   // stn[29].wipBtn[35,0] := 1000;
   // stn[29].wipBtn[35,1] := 1000;
   // stn[29].wipBtn[35,2] := 1000;
   // stn[29].wipBtn[35,3] := 1000;
   // stn[29].wipBtn[35,4] := 1000;
   // stn[29].wipBtn[35,5] := 1000;
   // stn[29].wipBtn[35,6] := 1000;
   // stn[29].wipBtn[35,7] := 1000;
   // stn[29].wipBtn[36,0] := 1000;
   // stn[29].wipBtn[36,1] := 1000;
   // stn[29].wipBtn[36,2] := 1000;
   // stn[29].wipBtn[36,3] := 1000;
   // stn[29].wipBtn[36,4] := 1000;
   // stn[29].wipBtn[36,5] := 1000;
   // stn[29].wipBtn[36,6] := 1000;
   // stn[29].wipBtn[36,7] := 1000;
   // stn[29].wipBtn[37,0] := 1000;
   // stn[29].wipBtn[37,1] := 1000;
   // stn[29].wipBtn[37,2] := 1000;
   // stn[29].wipBtn[37,3] := 1000;
   // stn[29].wipBtn[37,4] := 1000;
   // stn[29].wipBtn[37,5] := 1000;
   // stn[29].wipBtn[37,6] := 1000;
   // stn[29].wipBtn[37,7] := 1000;
   // stn[29].wipBtn[38,0] := 1000;
   // stn[29].wipBtn[38,1] := 1000;
   // stn[29].wipBtn[38,2] := 1000;
   // stn[29].wipBtn[38,3] := 1000;
   // stn[29].wipBtn[38,4] := 1000;
   // stn[29].wipBtn[38,5] := 1000;
   // stn[29].wipBtn[38,6] := 1000;
   // stn[29].wipBtn[38,7] := 1000;
   // stn[29].wipBtn[39,0] := 1000;
   // stn[29].wipBtn[39,1] := 1000;
   // stn[29].wipBtn[39,2] := 1000;
   // stn[29].wipBtn[39,3] := 1000;
   // stn[29].wipBtn[39,4] := 1000;
   // stn[29].wipBtn[39,5] := 1000;
   // stn[29].wipBtn[39,6] := 1000;
   // stn[29].wipBtn[39,7] := 1000;
   // stn[29].wipBtn[40,0] := 1000;
   // stn[29].wipBtn[40,1] := 1000;
   // stn[29].wipBtn[40,2] := 1000;
   // stn[29].wipBtn[40,3] := 1000;
   // stn[29].wipBtn[40,4] := 1000;
   // stn[29].wipBtn[40,5] := 1000;
   // stn[29].wipBtn[40,6] := 1000;
   // stn[29].wipBtn[40,7] := 1000;
   // stn[29].wipBtn[41,0] := 1000;
   // stn[29].wipBtn[41,1] := 1000;
   // stn[29].wipBtn[41,2] := 1000;
   // stn[29].wipBtn[41,3] := 1000;
   // stn[29].wipBtn[41,4] := 1000;
   // stn[29].wipBtn[41,5] := 1000;
   // stn[29].wipBtn[41,6] := 1000;
   // stn[29].wipBtn[41,7] := 1000;
   // stn[29].wipBtn[42,0] := 1000;
   // stn[29].wipBtn[42,1] := 1000;
   // stn[29].wipBtn[42,2] := 1000;
   // stn[29].wipBtn[42,3] := 1000;
   // stn[29].wipBtn[42,4] := 1000;
   // stn[29].wipBtn[42,5] := 1000;
   // stn[29].wipBtn[42,6] := 1000;
   // stn[29].wipBtn[42,7] := 1000;
   // stn[29].wipBtn[43,0] := 1000;
   // stn[29].wipBtn[43,1] := 1000;
   // stn[29].wipBtn[43,2] := 1000;
   // stn[29].wipBtn[43,3] := 1000;
   // stn[29].wipBtn[43,4] := 1000;
   // stn[29].wipBtn[43,5] := 1000;
   // stn[29].wipBtn[43,6] := 1000;
   // stn[29].wipBtn[43,7] := 1000;
   // stn[29].wipBtn[44,0] := 1000;
   // stn[29].wipBtn[44,1] := 1000;
   // stn[29].wipBtn[44,2] := 1000;
   // stn[29].wipBtn[44,3] := 1000;
   // stn[29].wipBtn[44,4] := 1000;
   // stn[29].wipBtn[44,5] := 1000;
   // stn[29].wipBtn[44,6] := 1000;
   // stn[29].wipBtn[44,7] := 1000;
   // stn[29].wipBtn[45,0] := 1000;
   // stn[29].wipBtn[45,1] := 1000;
   // stn[29].wipBtn[45,2] := 1000;
   // stn[29].wipBtn[45,3] := 1000;
   // stn[29].wipBtn[45,4] := 1000;
   // stn[29].wipBtn[45,5] := 1000;
   // stn[29].wipBtn[45,6] := 1000;
   // stn[29].wipBtn[45,7] := 1000;
   // stn[29].wipBtn[46,0] := 1000;
   // stn[29].wipBtn[46,1] := 1000;
   // stn[29].wipBtn[46,2] := 1000;
   // stn[29].wipBtn[46,3] := 1000;
   // stn[29].wipBtn[46,4] := 1000;
   // stn[29].wipBtn[46,5] := 1000;
   // stn[29].wipBtn[46,6] := 1000;
   // stn[29].wipBtn[46,7] := 1000;
   // stn[29].wipBtn[47,0] := 1000;
   // stn[29].wipBtn[47,1] := 1000;
   // stn[29].wipBtn[47,2] := 1000;
   // stn[29].wipBtn[47,3] := 1000;
   // stn[29].wipBtn[47,4] := 1000;
   // stn[29].wipBtn[47,5] := 1000;
   // stn[29].wipBtn[47,6] := 1000;
   // stn[29].wipBtn[47,7] := 1000;
   // stn[29].wipBtn[48,0] := 1000;
   // stn[29].wipBtn[48,1] := 1000;
   // stn[29].wipBtn[48,2] := 1000;
   // stn[29].wipBtn[48,3] := 1000;
   // stn[29].wipBtn[48,4] := 1000;
   // stn[29].wipBtn[48,5] := 1000;
   // stn[29].wipBtn[48,6] := 1000;
   // stn[29].wipBtn[48,7] := 1000;
   // stn[29].wipBtn[49,0] := 1000;
   // stn[29].wipBtn[49,1] := 1000;
   // stn[29].wipBtn[49,2] := 1000;
   // stn[29].wipBtn[49,3] := 1000;
   // stn[29].wipBtn[49,4] := 1000;
   // stn[29].wipBtn[49,5] := 1000;
   // stn[29].wipBtn[49,6] := 1000;
   // stn[29].wipBtn[49,7] := 1000;
   // stn[30].wipBtn[0,0] := 1000;
   // stn[30].wipBtn[0,1] := 1000;
   // stn[30].wipBtn[0,2] := 1000;
   // stn[30].wipBtn[0,3] := 1000;
   // stn[30].wipBtn[0,4] := 1000;
   // stn[30].wipBtn[0,5] := 1000;
   // stn[30].wipBtn[0,6] := 1000;
   // stn[30].wipBtn[0,7] := 57000;
   // stn[30].wipBtn[1,0] := 1000;
   // stn[30].wipBtn[1,1] := 1000;
   // stn[30].wipBtn[1,2] := 1000;
   // stn[30].wipBtn[1,3] := 1000;
   // stn[30].wipBtn[1,4] := 1000;
   // stn[30].wipBtn[1,5] := 1000;
   // stn[30].wipBtn[1,6] := 1000;
   // stn[30].wipBtn[1,7] := 1000;
   // stn[30].wipBtn[2,0] := 1000;
   // stn[30].wipBtn[2,1] := 1000;
   // stn[30].wipBtn[2,2] := 1000;
   // stn[30].wipBtn[2,3] := 1000;
   // stn[30].wipBtn[2,4] := 1000;
   // stn[30].wipBtn[2,5] := 1000;
   // stn[30].wipBtn[2,6] := 1000;
   // stn[30].wipBtn[2,7] := 1000;
   // stn[30].wipBtn[3,0] := 1000;
   // stn[30].wipBtn[3,1] := 1000;
   // stn[30].wipBtn[3,2] := 1000;
   // stn[30].wipBtn[3,3] := 1000;
   // stn[30].wipBtn[3,4] := 1000;
   // stn[30].wipBtn[3,5] := 1000;
   // stn[30].wipBtn[3,6] := 1000;
   // stn[30].wipBtn[3,7] := 1000;
   // stn[30].wipBtn[4,0] := 1000;
   // stn[30].wipBtn[4,1] := 1000;
   // stn[30].wipBtn[4,2] := 1000;
   // stn[30].wipBtn[4,3] := 1000;
   // stn[30].wipBtn[4,4] := 1000;
   // stn[30].wipBtn[4,5] := 1000;
   // stn[30].wipBtn[4,6] := 1000;
   // stn[30].wipBtn[4,7] := 1000;
   // stn[30].wipBtn[5,0] := 1000;
   // stn[30].wipBtn[5,1] := 1000;
   // stn[30].wipBtn[5,2] := 1000;
   // stn[30].wipBtn[5,3] := 1000;
   // stn[30].wipBtn[5,4] := 1000;
   // stn[30].wipBtn[5,5] := 1000;
   // stn[30].wipBtn[5,6] := 1000;
   // stn[30].wipBtn[5,7] := 1000;
   // stn[30].wipBtn[6,0] := 1000;
   // stn[30].wipBtn[6,1] := 1000;
   // stn[30].wipBtn[6,2] := 1000;
   // stn[30].wipBtn[6,3] := 1000;
   // stn[30].wipBtn[6,4] := 1000;
   // stn[30].wipBtn[6,5] := 1000;
   // stn[30].wipBtn[6,6] := 1000;
   // stn[30].wipBtn[6,7] := 1000;
   // stn[30].wipBtn[7,0] := 1000;
   // stn[30].wipBtn[7,1] := 1000;
   // stn[30].wipBtn[7,2] := 1000;
   // stn[30].wipBtn[7,3] := 1000;
   // stn[30].wipBtn[7,4] := 1000;
   // stn[30].wipBtn[7,5] := 1000;
   // stn[30].wipBtn[7,6] := 1000;
   // stn[30].wipBtn[7,7] := 1000;
   // stn[30].wipBtn[8,0] := 1000;
   // stn[30].wipBtn[8,1] := 1000;
   // stn[30].wipBtn[8,2] := 1000;
   // stn[30].wipBtn[8,3] := 1000;
   // stn[30].wipBtn[8,4] := 1000;
   // stn[30].wipBtn[8,5] := 1000;
   // stn[30].wipBtn[8,6] := 1000;
   // stn[30].wipBtn[8,7] := 1000;
   // stn[30].wipBtn[9,0] := 1000;
   // stn[30].wipBtn[9,1] := 1000;
   // stn[30].wipBtn[9,2] := 1000;
   // stn[30].wipBtn[9,3] := 1000;
   // stn[30].wipBtn[9,4] := 1000;
   // stn[30].wipBtn[9,5] := 1000;
   // stn[30].wipBtn[9,6] := 1000;
   // stn[30].wipBtn[9,7] := 1000;
   // stn[30].wipBtn[10,0] := 1000;
   // stn[30].wipBtn[10,1] := 1000;
   // stn[30].wipBtn[10,2] := 1000;
   // stn[30].wipBtn[10,3] := 1000;
   // stn[30].wipBtn[10,4] := 1000;
   // stn[30].wipBtn[10,5] := 1000;
   // stn[30].wipBtn[10,6] := 1000;
   // stn[30].wipBtn[10,7] := 1000;
   // stn[30].wipBtn[11,0] := 1000;
   // stn[30].wipBtn[11,1] := 1000;
   // stn[30].wipBtn[11,2] := 1000;
   // stn[30].wipBtn[11,3] := 1000;
   // stn[30].wipBtn[11,4] := 1000;
   // stn[30].wipBtn[11,5] := 1000;
   // stn[30].wipBtn[11,6] := 1000;
   // stn[30].wipBtn[11,7] := 1000;
   // stn[30].wipBtn[12,0] := 1000;
   // stn[30].wipBtn[12,1] := 1000;
   // stn[30].wipBtn[12,2] := 1000;
   // stn[30].wipBtn[12,3] := 1000;
   // stn[30].wipBtn[12,4] := 1000;
   // stn[30].wipBtn[12,5] := 1000;
   // stn[30].wipBtn[12,6] := 1000;
   // stn[30].wipBtn[12,7] := 1000;
   // stn[30].wipBtn[13,0] := 1000;
   // stn[30].wipBtn[13,1] := 1000;
   // stn[30].wipBtn[13,2] := 1000;
   // stn[30].wipBtn[13,3] := 1000;
   // stn[30].wipBtn[13,4] := 1000;
   // stn[30].wipBtn[13,5] := 1000;
   // stn[30].wipBtn[13,6] := 1000;
   // stn[30].wipBtn[13,7] := 1000;
   // stn[30].wipBtn[14,0] := 1000;
   // stn[30].wipBtn[14,1] := 1000;
   // stn[30].wipBtn[14,2] := 1000;
   // stn[30].wipBtn[14,3] := 1000;
   // stn[30].wipBtn[14,4] := 1000;
   // stn[30].wipBtn[14,5] := 1000;
   // stn[30].wipBtn[14,6] := 1000;
   // stn[30].wipBtn[14,7] := 1000;
   // stn[30].wipBtn[15,0] := 1000;
   // stn[30].wipBtn[15,1] := 1000;
   // stn[30].wipBtn[15,2] := 1000;
   // stn[30].wipBtn[15,3] := 1000;
   // stn[30].wipBtn[15,4] := 1000;
   // stn[30].wipBtn[15,5] := 1000;
   // stn[30].wipBtn[15,6] := 1000;
   // stn[30].wipBtn[15,7] := 1000;
   // stn[30].wipBtn[16,0] := 1000;
   // stn[30].wipBtn[16,1] := 1000;
   // stn[30].wipBtn[16,2] := 1000;
   // stn[30].wipBtn[16,3] := 1000;
   // stn[30].wipBtn[16,4] := 1000;
   // stn[30].wipBtn[16,5] := 1000;
   // stn[30].wipBtn[16,6] := 1000;
   // stn[30].wipBtn[16,7] := 1000;
   // stn[30].wipBtn[17,0] := 1000;
   // stn[30].wipBtn[17,1] := 1000;
   // stn[30].wipBtn[17,2] := 1000;
   // stn[30].wipBtn[17,3] := 1000;
   // stn[30].wipBtn[17,4] := 1000;
   // stn[30].wipBtn[17,5] := 1000;
   // stn[30].wipBtn[17,6] := 1000;
   // stn[30].wipBtn[17,7] := 1000;
   // stn[30].wipBtn[18,0] := 1000;
   // stn[30].wipBtn[18,1] := 1000;
   // stn[30].wipBtn[18,2] := 1000;
   // stn[30].wipBtn[18,3] := 1000;
   // stn[30].wipBtn[18,4] := 1000;
   // stn[30].wipBtn[18,5] := 1000;
   // stn[30].wipBtn[18,6] := 1000;
   // stn[30].wipBtn[18,7] := 1000;
   // stn[30].wipBtn[19,0] := 1000;
   // stn[30].wipBtn[19,1] := 1000;
   // stn[30].wipBtn[19,2] := 1000;
   // stn[30].wipBtn[19,3] := 1000;
   // stn[30].wipBtn[19,4] := 1000;
   // stn[30].wipBtn[19,5] := 1000;
   // stn[30].wipBtn[19,6] := 1000;
   // stn[30].wipBtn[19,7] := 1000;
   // stn[30].wipBtn[20,0] := 1000;
   // stn[30].wipBtn[20,1] := 1000;
   // stn[30].wipBtn[20,2] := 1000;
   // stn[30].wipBtn[20,3] := 1000;
   // stn[30].wipBtn[20,4] := 1000;
   // stn[30].wipBtn[20,5] := 1000;
   // stn[30].wipBtn[20,6] := 1000;
   // stn[30].wipBtn[20,7] := 1000;
   // stn[30].wipBtn[21,0] := 1000;
   // stn[30].wipBtn[21,1] := 1000;
   // stn[30].wipBtn[21,2] := 1000;
   // stn[30].wipBtn[21,3] := 1000;
   // stn[30].wipBtn[21,4] := 1000;
   // stn[30].wipBtn[21,5] := 1000;
   // stn[30].wipBtn[21,6] := 1000;
   // stn[30].wipBtn[21,7] := 1000;
   // stn[30].wipBtn[22,0] := 1000;
   // stn[30].wipBtn[22,1] := 1000;
   // stn[30].wipBtn[22,2] := 1000;
   // stn[30].wipBtn[22,3] := 1000;
   // stn[30].wipBtn[22,4] := 1000;
   // stn[30].wipBtn[22,5] := 1000;
   // stn[30].wipBtn[22,6] := 1000;
   // stn[30].wipBtn[22,7] := 1000;
   // stn[30].wipBtn[23,0] := 1000;
   // stn[30].wipBtn[23,1] := 1000;
   // stn[30].wipBtn[23,2] := 1000;
   // stn[30].wipBtn[23,3] := 1000;
   // stn[30].wipBtn[23,4] := 1000;
   // stn[30].wipBtn[23,5] := 1000;
   // stn[30].wipBtn[23,6] := 1000;
   // stn[30].wipBtn[23,7] := 1000;
   // stn[30].wipBtn[24,0] := 1000;
   // stn[30].wipBtn[24,1] := 1000;
   // stn[30].wipBtn[24,2] := 1000;
   // stn[30].wipBtn[24,3] := 1000;
   // stn[30].wipBtn[24,4] := 1000;
   // stn[30].wipBtn[24,5] := 1000;
   // stn[30].wipBtn[24,6] := 1000;
   // stn[30].wipBtn[24,7] := 1000;
   // stn[30].wipBtn[25,0] := 1000;
   // stn[30].wipBtn[25,1] := 1000;
   // stn[30].wipBtn[25,2] := 1000;
   // stn[30].wipBtn[25,3] := 1000;
   // stn[30].wipBtn[25,4] := 1000;
   // stn[30].wipBtn[25,5] := 1000;
   // stn[30].wipBtn[25,6] := 1000;
   // stn[30].wipBtn[25,7] := 1000;
   // stn[30].wipBtn[26,0] := 1000;
   // stn[30].wipBtn[26,1] := 1000;
   // stn[30].wipBtn[26,2] := 1000;
   // stn[30].wipBtn[26,3] := 1000;
   // stn[30].wipBtn[26,4] := 1000;
   // stn[30].wipBtn[26,5] := 1000;
   // stn[30].wipBtn[26,6] := 1000;
   // stn[30].wipBtn[26,7] := 1000;
   // stn[30].wipBtn[27,0] := 1000;
   // stn[30].wipBtn[27,1] := 1000;
   // stn[30].wipBtn[27,2] := 1000;
   // stn[30].wipBtn[27,3] := 1000;
   // stn[30].wipBtn[27,4] := 1000;
   // stn[30].wipBtn[27,5] := 1000;
   // stn[30].wipBtn[27,6] := 1000;
   // stn[30].wipBtn[27,7] := 1000;
   // stn[30].wipBtn[28,0] := 1000;
   // stn[30].wipBtn[28,1] := 1000;
   // stn[30].wipBtn[28,2] := 1000;
   // stn[30].wipBtn[28,3] := 1000;
   // stn[30].wipBtn[28,4] := 1000;
   // stn[30].wipBtn[28,5] := 1000;
   // stn[30].wipBtn[28,6] := 1000;
   // stn[30].wipBtn[28,7] := 1000;
   // stn[30].wipBtn[29,0] := 1000;
   // stn[30].wipBtn[29,1] := 1000;
   // stn[30].wipBtn[29,2] := 1000;
   // stn[30].wipBtn[29,3] := 1000;
   // stn[30].wipBtn[29,4] := 1000;
   // stn[30].wipBtn[29,5] := 1000;
   // stn[30].wipBtn[29,6] := 1000;
   // stn[30].wipBtn[29,7] := 1000;
   // stn[30].wipBtn[30,0] := 1000;
   // stn[30].wipBtn[30,1] := 1000;
   // stn[30].wipBtn[30,2] := 1000;
   // stn[30].wipBtn[30,3] := 1000;
   // stn[30].wipBtn[30,4] := 1000;
   // stn[30].wipBtn[30,5] := 1000;
   // stn[30].wipBtn[30,6] := 1000;
   // stn[30].wipBtn[30,7] := 1000;
   // stn[30].wipBtn[31,0] := 1000;
   // stn[30].wipBtn[31,1] := 1000;
   // stn[30].wipBtn[31,2] := 1000;
   // stn[30].wipBtn[31,3] := 1000;
   // stn[30].wipBtn[31,4] := 1000;
   // stn[30].wipBtn[31,5] := 1000;
   // stn[30].wipBtn[31,6] := 1000;
   // stn[30].wipBtn[31,7] := 1000;
   // stn[30].wipBtn[32,0] := 1000;
   // stn[30].wipBtn[32,1] := 1000;
   // stn[30].wipBtn[32,2] := 1000;
   // stn[30].wipBtn[32,3] := 1000;
   // stn[30].wipBtn[32,4] := 1000;
   // stn[30].wipBtn[32,5] := 1000;
   // stn[30].wipBtn[32,6] := 1000;
   // stn[30].wipBtn[32,7] := 1000;
   // stn[30].wipBtn[33,0] := 1000;
   // stn[30].wipBtn[33,1] := 1000;
   // stn[30].wipBtn[33,2] := 1000;
   // stn[30].wipBtn[33,3] := 1000;
   // stn[30].wipBtn[33,4] := 1000;
   // stn[30].wipBtn[33,5] := 1000;
   // stn[30].wipBtn[33,6] := 1000;
   // stn[30].wipBtn[33,7] := 1000;
   // stn[30].wipBtn[34,0] := 1000;
   // stn[30].wipBtn[34,1] := 1000;
   // stn[30].wipBtn[34,2] := 1000;
   // stn[30].wipBtn[34,3] := 1000;
   // stn[30].wipBtn[34,4] := 1000;
   // stn[30].wipBtn[34,5] := 1000;
   // stn[30].wipBtn[34,6] := 1000;
   // stn[30].wipBtn[34,7] := 1000;
   // stn[30].wipBtn[35,0] := 1000;
   // stn[30].wipBtn[35,1] := 1000;
   // stn[30].wipBtn[35,2] := 1000;
   // stn[30].wipBtn[35,3] := 1000;
   // stn[30].wipBtn[35,4] := 1000;
   // stn[30].wipBtn[35,5] := 1000;
   // stn[30].wipBtn[35,6] := 1000;
   // stn[30].wipBtn[35,7] := 1000;
   // stn[30].wipBtn[36,0] := 1000;
   // stn[30].wipBtn[36,1] := 1000;
   // stn[30].wipBtn[36,2] := 1000;
   // stn[30].wipBtn[36,3] := 1000;
   // stn[30].wipBtn[36,4] := 1000;
   // stn[30].wipBtn[36,5] := 1000;
   // stn[30].wipBtn[36,6] := 1000;
   // stn[30].wipBtn[36,7] := 1000;
   // stn[30].wipBtn[37,0] := 1000;
   // stn[30].wipBtn[37,1] := 1000;
   // stn[30].wipBtn[37,2] := 1000;
   // stn[30].wipBtn[37,3] := 1000;
   // stn[30].wipBtn[37,4] := 1000;
   // stn[30].wipBtn[37,5] := 1000;
   // stn[30].wipBtn[37,6] := 1000;
   // stn[30].wipBtn[37,7] := 1000;
   // stn[30].wipBtn[38,0] := 1000;
   // stn[30].wipBtn[38,1] := 1000;
   // stn[30].wipBtn[38,2] := 1000;
   // stn[30].wipBtn[38,3] := 1000;
   // stn[30].wipBtn[38,4] := 1000;
   // stn[30].wipBtn[38,5] := 1000;
   // stn[30].wipBtn[38,6] := 1000;
   // stn[30].wipBtn[38,7] := 1000;
   // stn[30].wipBtn[39,0] := 1000;
   // stn[30].wipBtn[39,1] := 1000;
   // stn[30].wipBtn[39,2] := 1000;
   // stn[30].wipBtn[39,3] := 1000;
   // stn[30].wipBtn[39,4] := 1000;
   // stn[30].wipBtn[39,5] := 1000;
   // stn[30].wipBtn[39,6] := 1000;
   // stn[30].wipBtn[39,7] := 1000;
   // stn[30].wipBtn[40,0] := 1000;
   // stn[30].wipBtn[40,1] := 1000;
   // stn[30].wipBtn[40,2] := 1000;
   // stn[30].wipBtn[40,3] := 1000;
   // stn[30].wipBtn[40,4] := 1000;
   // stn[30].wipBtn[40,5] := 1000;
   // stn[30].wipBtn[40,6] := 1000;
   // stn[30].wipBtn[40,7] := 1000;
   // stn[30].wipBtn[41,0] := 1000;
   // stn[30].wipBtn[41,1] := 1000;
   // stn[30].wipBtn[41,2] := 1000;
   // stn[30].wipBtn[41,3] := 1000;
   // stn[30].wipBtn[41,4] := 1000;
   // stn[30].wipBtn[41,5] := 1000;
   // stn[30].wipBtn[41,6] := 1000;
   // stn[30].wipBtn[41,7] := 1000;
   // stn[30].wipBtn[42,0] := 1000;
   // stn[30].wipBtn[42,1] := 1000;
   // stn[30].wipBtn[42,2] := 1000;
   // stn[30].wipBtn[42,3] := 1000;
   // stn[30].wipBtn[42,4] := 1000;
   // stn[30].wipBtn[42,5] := 1000;
   // stn[30].wipBtn[42,6] := 1000;
   // stn[30].wipBtn[42,7] := 1000;
   // stn[30].wipBtn[43,0] := 1000;
   // stn[30].wipBtn[43,1] := 1000;
   // stn[30].wipBtn[43,2] := 1000;
   // stn[30].wipBtn[43,3] := 1000;
   // stn[30].wipBtn[43,4] := 1000;
   // stn[30].wipBtn[43,5] := 1000;
   // stn[30].wipBtn[43,6] := 1000;
   // stn[30].wipBtn[43,7] := 1000;
   // stn[30].wipBtn[44,0] := 1000;
   // stn[30].wipBtn[44,1] := 1000;
   // stn[30].wipBtn[44,2] := 1000;
   // stn[30].wipBtn[44,3] := 1000;
   // stn[30].wipBtn[44,4] := 1000;
   // stn[30].wipBtn[44,5] := 1000;
   // stn[30].wipBtn[44,6] := 1000;
   // stn[30].wipBtn[44,7] := 1000;
   // stn[30].wipBtn[45,0] := 1000;
   // stn[30].wipBtn[45,1] := 1000;
   // stn[30].wipBtn[45,2] := 1000;
   // stn[30].wipBtn[45,3] := 1000;
   // stn[30].wipBtn[45,4] := 1000;
   // stn[30].wipBtn[45,5] := 1000;
   // stn[30].wipBtn[45,6] := 1000;
   // stn[30].wipBtn[45,7] := 1000;
   // stn[30].wipBtn[46,0] := 1000;
   // stn[30].wipBtn[46,1] := 1000;
   // stn[30].wipBtn[46,2] := 1000;
   // stn[30].wipBtn[46,3] := 1000;
   // stn[30].wipBtn[46,4] := 1000;
   // stn[30].wipBtn[46,5] := 1000;
   // stn[30].wipBtn[46,6] := 1000;
   // stn[30].wipBtn[46,7] := 1000;
   // stn[30].wipBtn[47,0] := 1000;
   // stn[30].wipBtn[47,1] := 1000;
   // stn[30].wipBtn[47,2] := 1000;
   // stn[30].wipBtn[47,3] := 1000;
   // stn[30].wipBtn[47,4] := 1000;
   // stn[30].wipBtn[47,5] := 1000;
   // stn[30].wipBtn[47,6] := 1000;
   // stn[30].wipBtn[47,7] := 1000;
   // stn[30].wipBtn[48,0] := 1000;
   // stn[30].wipBtn[48,1] := 1000;
   // stn[30].wipBtn[48,2] := 1000;
   // stn[30].wipBtn[48,3] := 1000;
   // stn[30].wipBtn[48,4] := 1000;
   // stn[30].wipBtn[48,5] := 1000;
   // stn[30].wipBtn[48,6] := 1000;
   // stn[30].wipBtn[48,7] := 1000;
   // stn[30].wipBtn[49,0] := 1000;
   // stn[30].wipBtn[49,1] := 1000;
   // stn[30].wipBtn[49,2] := 1000;
   // stn[30].wipBtn[49,3] := 1000;
   // stn[30].wipBtn[49,4] := 1000;
   // stn[30].wipBtn[49,5] := 1000;
   // stn[30].wipBtn[49,6] := 1000;
   // stn[30].wipBtn[49,7] := 1000;
END_TYPE

TYPE "Recipe: PN Text"
VERSION : 0.1
   STRUCT
      pnText : Array[0.."pnLibCount"] of WString["sStringLen"];
   END_STRUCT;
END_TYPE

// folder: KP8

TYPE "KP8 Driver: Parameters: 1 Button"
   STRUCT
      activate : Bool;   // true = button on, flase = button off
      cOn1 : String[10];   // color when button is in pressed state. valid entries: 'red', 'green', 'blue', 'yellow', 'white', 'off'
      cOn2 : String[10];   // second flash color when button is pressed and flashing is enabled. valid entries: 'red', 'green', 'blue', 'yellow', 'white', 'off'
      cOff : String[10];   // color when button is in un-pressed state. valid entries: 'red', 'green', 'blue', 'yellow', 'white', 'off'
      flash : Bool;   // false = color 1, true = color 2. set to clock bit to flash at that rate
      group : Int;   // 0 disables. buttons in groups have a mutually exclusive 'on' state.
      mode : Bool;   // true = maintained, fales = momentary
   END_STRUCT;
END_TYPE

TYPE "KP8 Driver: Button States"
   STRUCT
      btn : Array[0..7] of Bool;
   END_STRUCT;
END_TYPE

TYPE "KP8 Driver: Parameters: 8 Buttons"
   STRUCT
      btn : Array[0..7] of "KP8 Driver: Parameters: 1 Button";
   END_STRUCT;
END_TYPE

TYPE "KP8 Driver: Feedback Data"
   STRUCT
      acutal : "KP8 Driver: Button States";
      falling : "KP8 Driver: Button States";
      rising : "KP8 Driver: Button States";
   END_STRUCT;
END_TYPE

// folder: Main HMI

TYPE "Part Call Screen"
   STRUCT
      row : Array[0.."partReqHmiRowCount"] of "Table Row";
   END_STRUCT;
END_TYPE

TYPE "Table Row"
   STRUCT
      address : UInt;
      ordered : Bool;
      pbSelection : Struct
         actuate : Bool;
         animate : USInt;
      END_STRUCT;
      rtBackground : Struct
         animate : USInt;
      END_STRUCT;
      tfDropZone : Struct
         animate : USInt;
         value : WString[20];
      END_STRUCT;
      tfLine : Struct
         animate : USInt;
         value : WString[20];
      END_STRUCT;
      tfPartNumber : Struct
         animateDL : USInt;
         animateSL : USInt;
         value : WString[40];
      END_STRUCT;
      tfTime : Struct
         animate : USInt;
         value : WString[20];
      END_STRUCT;
   END_STRUCT;
END_TYPE

TYPE "Part Request Data"
   STRUCT
      row : Array[0.."partReqDataRowCount"] of "Table Row";
   END_STRUCT;
END_TYPE

TYPE "PB Data: Graphic/Text List"
   STRUCT
      actuate : Bool;
      animate : USInt;
      listSelect : UInt;
   END_STRUCT;
END_TYPE

TYPE "LED Sign Data"
   STRUCT
      row : Array[0.."ledRowCount"] of "Table Row";
   END_STRUCT;
END_TYPE

TYPE "PB Data: Text Label"
   STRUCT
      actuate : Bool;
      animate : USInt;
      label : WString[20];
   END_STRUCT;
END_TYPE

TYPE "IO Field Data: Part Number"
   STRUCT
      animate : USInt;
      inputFinished : Bool;
      value : WString[40];
   END_STRUCT;
END_TYPE

TYPE "Line Label Data"
   STRUCT
      animate : Struct
         bg : USInt;
         ioField : USInt;
      END_STRUCT;
      inputFinished : Bool;
      value : WString[10];
   END_STRUCT;
END_TYPE

TYPE "Drop Zone Data"
   STRUCT
      animate : Struct
         bg : USInt;
         ioField : USInt;
      END_STRUCT;
      inputFinished : Bool;
      value : WString[10];
   END_STRUCT;
END_TYPE

TYPE "IO Field Data: Timers"
   STRUCT
      animate : USInt;
      inputFinished : Bool;
      value : WString[5];
   END_STRUCT;
END_TYPE

TYPE "Table Nav: HMI"
   STRUCT
      top : "PB Data: Graphic/Text List";
      pageUp : "PB Data: Graphic/Text List";
      lineUp : "PB Data: Graphic/Text List";
      lineDown : "PB Data: Graphic/Text List";
      pageDown : "PB Data: Graphic/Text List";
      bottom : "PB Data: Graphic/Text List";
   END_STRUCT;
END_TYPE

TYPE "Simulated Stations"
   STRUCT
      down : "PB Data: Graphic/Text List";
      firstStn : Int;
      me : Array[0.."simKP8Count"] of "Station: Sim Data";
      up : "PB Data: Graphic/Text List";
   END_STRUCT;
END_TYPE

TYPE "Network Health Screen"
   STRUCT
      et200spPopUp : "Station: ET200SP Comm Debug Data";
      kp8PopUp : "Station: KP8 Comm Debug Data";
      pnioDevices : Array[1.."pnioDeviceCount"] of "PB Data: Text Label";
      selectedDevice : Int;
   END_STRUCT;
   // // pnioDevices[1] : volvo1601kp8
   // // pnioDevices[2] : volvo1601et200sp
   // // pnioDevices[3] : volvo1602kp8
   // // pnioDevices[4] : volvo1602et200sp
   // // pnioDevices[5] : volvo1603kp8
   // // pnioDevices[6] : volvo1603et200sp
   // // pnioDevices[7] : volvo1604kp8
   // // pnioDevices[8] : volvo1604et200sp
   // // pnioDevices[9] : volvo1605kp8
   // // pnioDevices[10] : volvo1605et200sp
   // // pnioDevices[11] : volvo1606kp8
   // // pnioDevices[12] : volvo1606et200sp
   // // pnioDevices[13] : volvo1607kp8
   // // pnioDevices[14] : volvo1607et200sp
   // // pnioDevices[15] : volvo1608kp8
   // // pnioDevices[16] : volvo1608et200sp
   // // pnioDevices[17] : volvo1609kp8
   // // pnioDevices[18] : volvo1609et200sp
   // // pnioDevices[19] : volvo1610kp8
   // // pnioDevices[20] : volvo1610et200sp
   // // pnioDevices[21] : volvo1611kp8
   // // pnioDevices[22] : volvo1611et200sp
   // // pnioDevices[23] : chm01kp8
   // // pnioDevices[24] : chm01et200sp
   // // pnioDevices[25] : chm02kp8
   // // pnioDevices[26] : chm02et200sp
   // // pnioDevices[27] : chm03kp8
   // // pnioDevices[28] : chm03et200sp
   // // pnioDevices[29] : chm04kp8
   // // pnioDevices[30] : chm04et200sp
   // // pnioDevices[31] : chm05kp8
   // // pnioDevices[32] : chm05et200sp
   // // pnioDevices[33] : cd001kp8
   // // pnioDevices[34] : cd001et200sp
   // // pnioDevices[35] : cd002kp8
   // // pnioDevices[36] : cd002et200sp
   // // pnioDevices[37] : cd003kp8
   // // pnioDevices[38] : cd003et200sp
   // // pnioDevices[39] : bfl01kp8
   // // pnioDevices[40] : bfl01et200sp
   // // pnioDevices[41] : bfl02kp8
   // // pnioDevices[42] : bfl02et200sp
   // // pnioDevices[43] : bfl03kp8
   // // pnioDevices[44] : bfl03et200sp
   // // pnioDevices[45] : lgs01kp8
   // // pnioDevices[46] : lgs01et200sp
   // // pnioDevices[47] : lgs02kp8
   // // pnioDevices[48] : lgs02et200sp
END_TYPE

TYPE "Table Nav: PLC"
   STRUCT
      top : Bool;
      pageUp : Bool;
      lineUp : Bool;
      lineDown : Bool;
      pageDown : Bool;
      bottom : Bool;
   END_STRUCT;
END_TYPE

// folder: Main HMI/Barcode

TYPE "Barcode Screen"
   STRUCT
      partNumber : WString[40];
      barcode : String;
      acknowledged : Bool;
      ordered : Bool;
   END_STRUCT;
END_TYPE

// folder: Main HMI/Settings Screen

TYPE "Settings"
   STRUCT
      alotted : "Settings Alotted";
      critical : "Settings Critical";
      kp8 : "Settings KP8";
      stations : "Settings Stations";
      partNumber : "Settings Part Number";
      viewingStation : "Settings Viewing Stations";
   END_STRUCT;
END_TYPE

TYPE "Settings Alotted"
   STRUCT
      assign : "PB Data: Text Label";
      ioField : "IO Field Data: Timers";
   END_STRUCT;
END_TYPE

TYPE "Settings Critical"
   STRUCT
      assign : "PB Data: Text Label";
      ioField : "IO Field Data: Timers";
   END_STRUCT;
END_TYPE

TYPE "Settings KP8"
   STRUCT
      selectButtons : "PB Data: Text Label";
      btnSelState : Array[0.."btnCount"] of Bool;
      buttons : Array[0.."btnCount"] of "PB Data: Text Label";
      selBtnNumber : Int;
      selCount : Int;
   END_STRUCT;
END_TYPE

TYPE "Settings Stations"
   STRUCT
      selectAll : "PB Data: Text Label";
      nextGroup : "PB Data: Graphic/Text List";
      prevGroup : "PB Data: Graphic/Text List";
      selectBtns : Array[0.."hmiSelStnCount"] of "PB Data: Text Label";
      selCount : Int;
      selNumber : Int;
   END_STRUCT;
END_TYPE

TYPE "Settings Part Number"
   STRUCT
      assign : "PB Data: Text Label";
      ioField : "IO Field Data: Part Number";
   END_STRUCT;
END_TYPE

TYPE "Settings Viewing Stations"
   STRUCT
      btns : Array[0.."btnCount"] of "Station: Assignment: Button Details";
      dzData : "Drop Zone Data";
      lineData : "Line Label Data";
      next : "PB Data: Graphic/Text List";
      previous : "PB Data: Graphic/Text List";
      "name" : WString[20];
   END_STRUCT;
END_TYPE

// folder: Recipe System

TYPE "Recipe: Wip"
   STRUCT
      dropZone : USInt;
      kp8Output : DWord;
      kp8LogicalState0 : Bool;
      kp8LogicalState1 : Bool;
      kp8LogicalState2 : Bool;
      kp8LogicalState3 : Bool;
      kp8LogicalState4 : Bool;
      kp8LogicalState5 : Bool;
      kp8LogicalState6 : Bool;
      kp8LogicalState7 : Bool;
      lineName : USInt;
      pnCode : DInt;
      stackLight : DWord;
      wipName : WString;
      wipNumber : UInt;
   END_STRUCT;
END_TYPE

TYPE "Recipe: Station"
   STRUCT
      wip : Array[0.."wipCount"] of "Recipe: Wip";
   END_STRUCT;
END_TYPE

// folder: Station

TYPE "Station: All Stations"
   STRUCT
      stn : Array[0.."stnCount"] of "Station: Single Station";
   END_STRUCT;
END_TYPE

TYPE "Station: Order States"
   STRUCT
      btn : Array[0.."btnCount"] of Int;
   END_STRUCT;
END_TYPE

TYPE "Station: KP8 Config"
VERSION : 0.1
   STRUCT
      activate : Bool;
      colorOn1 : String[10];
      colorOn2 : String[10];
      colorOff : String[10];
      flash : Bool;
      group : Int;
      mode : Bool;
   END_STRUCT;
END_TYPE

TYPE "Station: PN Code"
   STRUCT
      btn : Array[0.."btnCount"] of DInt;
   END_STRUCT;
END_TYPE

TYPE "Station: Single Station"
   STRUCT
      animate : Array[0.."btnCount"] of UInt;
      id : "Station: Id";
      ioData : "Station I/O Data";
      flags : "Station: Flags";
      kp8Config : "KP8 Driver: Parameters: 8 Buttons";
      kp8Logical : "KP8 Driver: Feedback Data";
      kp8Physical : "KP8 Driver: Feedback Data";
      orderState : Array[0.."btnCount"] of Int;
      pnCode : Array[0.."btnCount"] of DInt;
      timers : "Station: Timers";
      wipData : "Station: Loaded WIP Data";
   END_STRUCT;
END_TYPE

TYPE "Station: Animations"
   STRUCT
      btn : Array[0.."btnCount"] of UInt;
   END_STRUCT;
END_TYPE

TYPE "Station: Flags"
   STRUCT
      inSettingsScreen : Bool;
      newPN : Bool;
      pnGood : Array[0.."btnCount"] of Bool;
      resetStation : Bool;
      resetTimer : Array[0.."btnCount"] of Bool;
      stateTransition : Array[0.."btnCount"] of Bool;
   END_STRUCT;
END_TYPE

TYPE "Station: Timers"
   STRUCT
      elapsed : Array[0.."btnCount"] of Real;
      ptAllotted : Array[0.."btnCount"] of Real;
      ptCritical : Array[0.."btnCount"] of Real;
      remaining : Array[0.."btnCount"] of Real;
   END_STRUCT;
END_TYPE

TYPE "Station: Id"
   STRUCT
      dropZone : USInt;
      lineName : WString["sStringLen"];
   END_STRUCT;
END_TYPE

TYPE "Station: Loaded WIP Data"
   STRUCT
      number : UInt;
      "name" : WString["lStringLen"];
   END_STRUCT;
END_TYPE

// folder: Station/ET200SP

TYPE "ET200SP: IM Data"
   STRUCT
      bg : USInt;
      error : USInt;
      lnk01 : USInt;
      lnk02 : USInt;
      maint : USInt;
      pwr : USInt;
      run : USInt;
   END_STRUCT;
END_TYPE

TYPE "ET200SP: DQ Data"
   STRUCT
      bg : USInt;
      bgTem : USInt;
      diag : USInt;
      pwr : USInt;
      x0 : USInt;
      x1 : USInt;
      x2 : USInt;
      x3 : USInt;
      x4 : USInt;
      x5 : USInt;
      x6 : USInt;
      x7 : USInt;
   END_STRUCT;
END_TYPE

TYPE "ET200SP: Server Module Data"
   STRUCT
      bg : USInt;
   END_STRUCT;
END_TYPE

// folder: Station/Faceplate

TYPE "Station: Assignment: Button Details"
   STRUCT
      alloted : Struct
         animate : USInt;
         value : WString[10];
      END_STRUCT;
      critical : Struct
         animate : USInt;
         value : WString[10];
      END_STRUCT;
      label : Struct
         animate : USInt;
         value : WString[2];
      END_STRUCT;
      partNumber : Struct
         animate : USInt;
         value : WString[40];
      END_STRUCT;
      select : Struct
         actuate : Bool;
         animate : USInt;
      END_STRUCT;
   END_STRUCT;
END_TYPE

TYPE "Station: Sim Data"
   STRUCT
      stn : Struct
         animate : USInt;
         label : WString[20];
      END_STRUCT;
      btn : Struct
         actuate : Byte;
         animate : Array[0..7] of USInt;
         labels : Array[0..7] of WString [4];
      END_STRUCT;
   END_STRUCT;
END_TYPE

TYPE "Station: ET200SP Comm Debug Data"
   STRUCT
      dismissPB : Bool;
      IM : "ET200SP: IM Data";
      DQ01 : "ET200SP: DQ Data";
      DQ02 : "ET200SP: DQ Data";
      DQ03 : "ET200SP: DQ Data";
      profinetName : Struct
         animate : USInt;
         label : WString[20];
      END_STRUCT;
      serverModule : "ET200SP: Server Module Data";
   END_STRUCT;
END_TYPE

TYPE "Station: KP8 Comm Debug Data"
   STRUCT
      dismissPB : Bool;
      profinetName : Struct
         animate : USInt;
         label : WString[20];
      END_STRUCT;
      stencilBackground : USInt;
      X1P1 : Struct
         transmit : USInt;
         receive : USInt;
      END_STRUCT;
      X1P2 : Struct
         transmit : USInt;
         receive : USInt;
      END_STRUCT;
   END_STRUCT;
END_TYPE

// folder: Station/HMI Station

TYPE "HMIS: Part Selection Screen"
   STRUCT
      animate : Array[0.."hmiStnPartSelScrnBtnCnt"] of Int;
      pbs : DWord;
      txt : Array[0.."hmiStnPartSelScrnBtnCnt"] of WString [40];
   END_STRUCT;
END_TYPE

TYPE "HMIS: Compressed"
   STRUCT
      scrnSlctPrt : "HMIS: Part Selection Screen";
      scrnSlctMn : "HMIS: Menu Selection Screen";
      scrnTmplt : "HMIS: Template Screen";
   END_STRUCT;
END_TYPE

TYPE "HMIS: Menu Selection Screen"
   STRUCT
      animate : Array[0.."hmiStnMenuSelScrnBtnCnt"] of Int;
      pbs : DWord;
      txt : Array[0.."hmiStnMenuSelLblCnt"] of WString ["lStringLen"];
   END_STRUCT;
END_TYPE

TYPE "HMIS: Template Screen"
   STRUCT
      animate : Array[0.."hmiStnTmpltBtnCnt"] of Int;
      pb : DWord;
      text : Array[0.."hmiStnTmpltBtnCnt"] of WString ["lStringLen"];
   END_STRUCT;
END_TYPE

// folder: Station/KP8

TYPE "KP8 I/O Data"
   STRUCT
      input : Word;
      output : DWord;
   END_STRUCT;
END_TYPE

TYPE "Station I/O Data"
   STRUCT
      kp8 : "KP8 I/O Data";
      stkLight : DWord;
   END_STRUCT;
END_TYPE

// folder: (top level)

DATA_BLOCK "Debug"   // DB7
{ S7_Optimized_Access := 'TRUE' }
VERSION : 0.1
   VAR
      test : Bool;
      address : UInt;
      stn : Int;
      btn : Int;
   END_VAR
BEGIN
END_DATA_BLOCK

// folder: Global Data

DATA_BLOCK "EMP IDB"   // DB1
{ S7_Optimized_Access := 'TRUE' }
VERSION : 0.1
// stored: InstanceOfName EMP
"EMP"
BEGIN
END_DATA_BLOCK

